(* Logix 5000 project; controller Seperator 1756-L85E rev 33.11; software revision 33.01; part 5 of 7 *)
(* tags used below, declared in another part *)
   batchstrng : STRING;
   bottle_clamp_out_delay : TIMER;
   bottle_clamp_out_delayF1 : TIMER;
   CAP_clamps_out_Delay : TIMER;
   Capper_Head_Sequencer : DINT;
   colours : STRING[3];
   Filler_Index_complete : BOOL;
   Filling : SFC_STEP;
   Filling_Nozzle_Down_Delay1 : TIMER;
   Filling_Nozzle_up_Delay1 : TIMER;
   Logix_Status : Logix_Status_FP;
   Qtr_Sec_PLs : TIMER;
   Random : AOI_SIM_RNG_Simple;

PROGRAM Capper_Heads   (* main routine Initialisation *)
VAR
   Alias_Head_Clamp_Pressure_SP : ALIAS FOR Head_Clamp_Pressure_SP;
   Bottle_Clamp_Pressure_actual : REAL := 10.799999;
   Cap_Pressure : REAL := 9.4;
   Head1_98_Percent_temperatureSP : REAL := 176.4;
   Head_Clamp_Pressure_SP : REAL := 90.0;
   Head_Down : BOOL;
   Head_Down_Stage1 : REAL := 18.0;
   Head_Down_Stage2 : REAL := 27.0;
   Head_Injection_Pressure_SP : REAL := 75.0;
   Head_Injection_Stage1 : REAL := 18.75;
   Head_Injection_Stage2 : REAL := 33.75;
   Head_Injector_out_delay : TIMER := (PRE := 2000);
   Head_moving_Down : BOOL := 1;
   Head_moving_Up : BOOL;
   Head_Up : BOOL;
   Head_up_delay : TIMER := (PRE := 2000);
   Pump_Running : BOOL := 1;
   Rotary_Moulder_Head_Name : STRING := 'Head 1'; {constant, access None}
   ScratchPad1 : REAL := 0.9;
   ScratchPad2 : REAL := 0.9;
   ScratchPad3 : REAL := 0.75;
   ScratchPad4 : REAL := 0.75;
   ScratchPad5 : REAL := 3.6;
   ScratchPad6 : REAL;
END_VAR

ROUTINE Head_Control   (* ladder *)
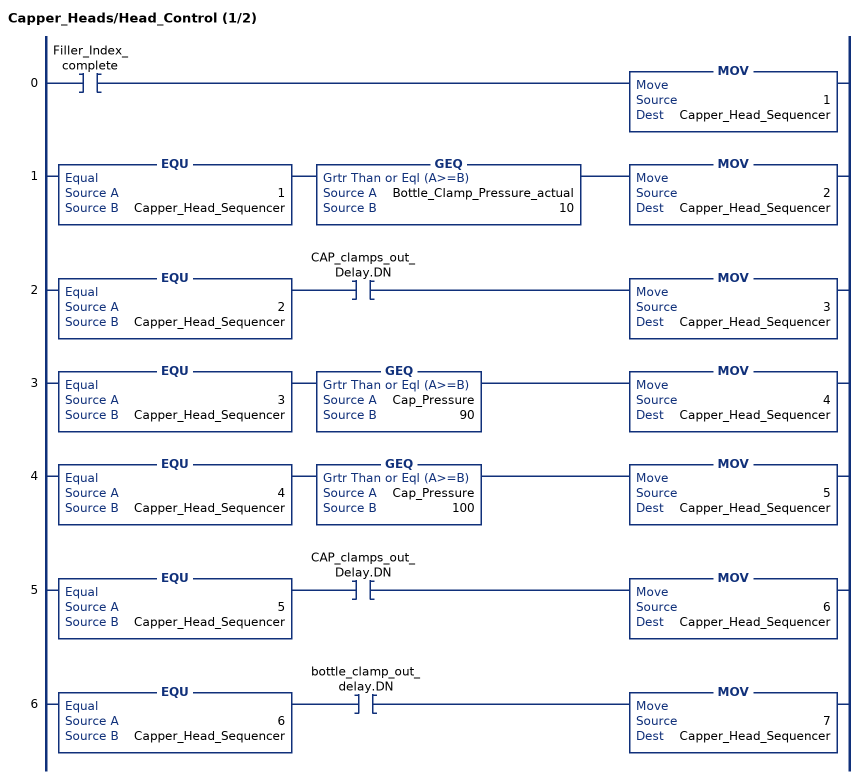
   0: XIC(Filler_Index_complete)MOV(1,Capper_Head_Sequencer);
   1: EQU(1,Capper_Head_Sequencer)GEQ(Bottle_Clamp_Pressure_actual,10)MOV(2,Capper_Head_Sequencer);
   2: EQU(2,Capper_Head_Sequencer)XIC(CAP_clamps_out_Delay.DN)MOV(3,Capper_Head_Sequencer);
   3: EQU(3,Capper_Head_Sequencer)GEQ(Cap_Pressure,90)MOV(4,Capper_Head_Sequencer);
   4: EQU(4,Capper_Head_Sequencer)GEQ(Cap_Pressure,100)MOV(5,Capper_Head_Sequencer);
   5: EQU(5,Capper_Head_Sequencer)XIC(CAP_clamps_out_Delay.DN)MOV(6,Capper_Head_Sequencer);
   6: EQU(6,Capper_Head_Sequencer)XIC(bottle_clamp_out_delay.DN)MOV(7,Capper_Head_Sequencer);
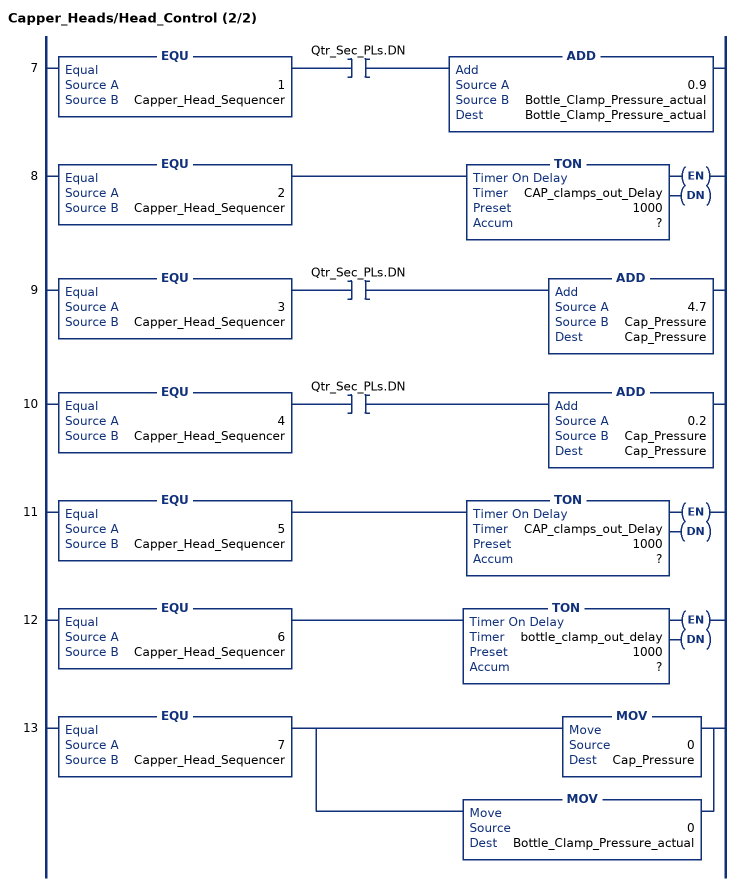
   7: EQU(1,Capper_Head_Sequencer)XIC(Qtr_Sec_PLs.DN)ADD(0.9,Bottle_Clamp_Pressure_actual,Bottle_Clamp_Pressure_actual);
   8: EQU(2,Capper_Head_Sequencer)TON(CAP_clamps_out_Delay,?,?);
   9: EQU(3,Capper_Head_Sequencer)XIC(Qtr_Sec_PLs.DN)ADD(4.7,Cap_Pressure,Cap_Pressure);
   10: EQU(4,Capper_Head_Sequencer)XIC(Qtr_Sec_PLs.DN)ADD(0.2,Cap_Pressure,Cap_Pressure);
   11: EQU(5,Capper_Head_Sequencer)TON(CAP_clamps_out_Delay,?,?);
   12: EQU(6,Capper_Head_Sequencer)TON(bottle_clamp_out_delay,?,?);
   13: EQU(7,Capper_Head_Sequencer)[MOV(0,Cap_Pressure) ,MOV(0,Bottle_Clamp_Pressure_actual) ];
END_ROUTINE

ROUTINE Head_HMI_Collation   (* ladder *)
END_ROUTINE

ROUTINE Initialisation   (* ladder *)
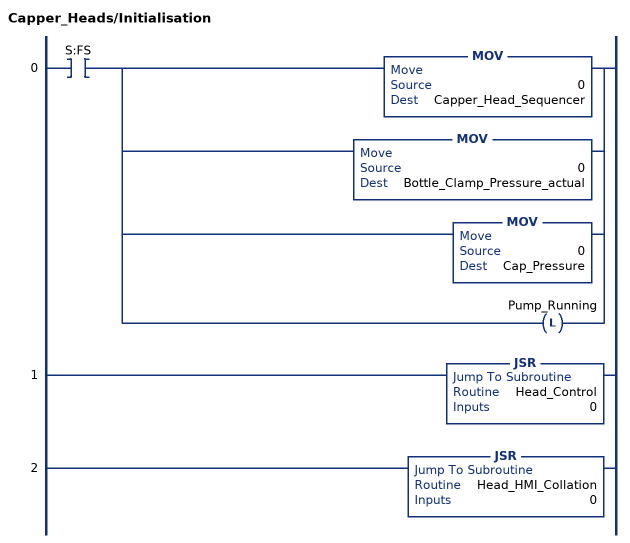
   0: XIC(S:FS)[MOV(0,Capper_Head_Sequencer) ,MOV(0,Bottle_Clamp_Pressure_actual) ,MOV(0,Cap_Pressure) ,OTL(Pump_Running) ];
   1: JSR(Head_Control,0);
   2: JSR(Head_HMI_Collation,0);
END_ROUTINE
END_PROGRAM

PROGRAM Controller_Fault   (* main routine Major_Controller_Fault *)

ROUTINE Major_Controller_Fault   (* ladder *)
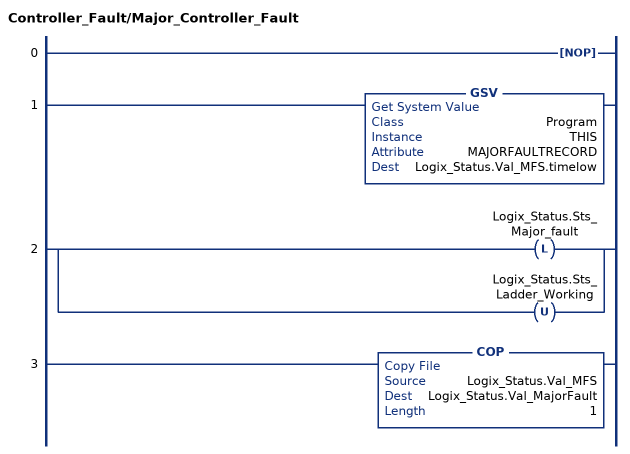
   0: NOP();
   1: GSV(Program,THIS,MAJORFAULTRECORD,Logix_Status.Val_MFS.timelow);
   2: [OTL(Logix_Status.Sts_Major_fault) ,OTU(Logix_Status.Sts_Ladder_Working) ];
   3: COP(Logix_Status.Val_MFS,Logix_Status.Val_MajorFault,1);
END_ROUTINE
END_PROGRAM

PROGRAM Filler   (* main routine Initialisation *)
VAR
   autoreset : TIMER := (PRE := 38913);
   autoresetpulse : BOOL;
   batchcountbase : DINT := 35000;
   batchcounter : DINT := 704;
   colourcounter : DINT := 2;
   Filler1_Heater_Tripped : ALARM_DIGITAL;
   Filler1_Hyd_Oil_Pressure_Low : ALARM_DIGITAL;
   Filler1_Hyd_Pump_Failure : ALARM_DIGITAL;
   Filler1_Index_Failure : ALARM_DIGITAL;
   Filler1_Overload : ALARM_DIGITAL;
   Filler_Efficiency_FTAE : BOOL[32];
   Filler_Fault_FTAE : BOOL[32];
   Filler_Heater_Tripped : BOOL;
   Filler_Hyd_Oil_Pressure_Low : BOOL;
   Filler_Hyd_Pump_Failure : BOOL;
   Filler_Index_Failure : BOOL;
   Filler_Overload : BOOL;
   Filler_Running : BOOL := 1;
   Filler_Warning_FTAE : BOOL[32];
   Index_Move : BOOL;
   Index_Move_Timer : TIMER := (PRE := 1000);
   m_slowperc_lim : REAL := 0.92;
   MetricsData : mtrcsdt := (PartId := 'Corner block', IdealCT := 23.7, GoodParts := 30066, ScrapParts := 5250, TotalParts := 35316, Running := 1, Monitored_Availability := 1, Machine_State := 1, BatchID := 'Batch ID 35704', Colour := 'White');
   mset_badperc : REAL := 0.07;   // Bad percentage valid: 1.0 - mset_goodperc
   mset_fltfudge : REAL := 0.93;   // fault distribution fudge factor do not change
   mset_fltoffset : DINT := 2;   // fault distribution offset do not change
   mset_goodperc : REAL := 0.85;   // Good percentage valid: 0.51 - 0.99
   mset_wrnfudge : REAL := 0.02;   // warning distribution fudge factor do not change
   mset_wrnoffset : DINT := 2;   // warning distribution offset do not change
   oneshots : DINT;
   tempDINT : DINT := 16;
   tempstring : STRING := '35704';
END_VAR

ROUTINE Filler_Alarms   (* ladder *)
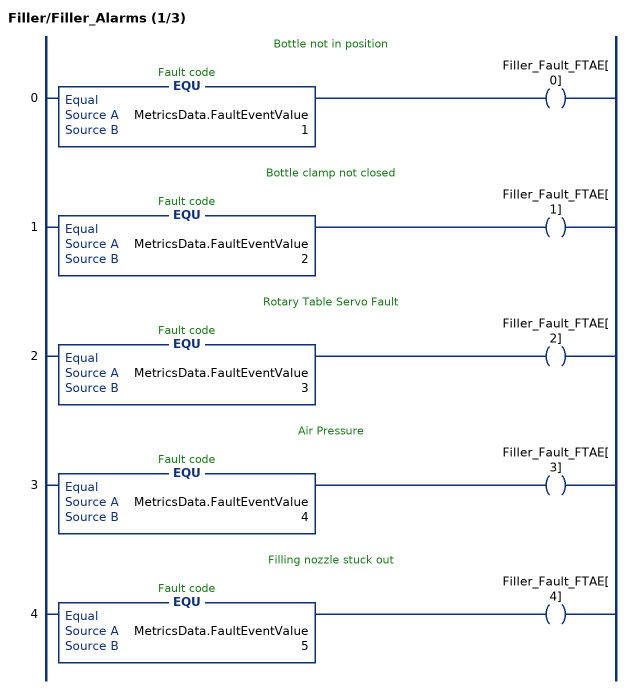
   // Bottle not in position
   0: EQU(MetricsData.FaultEventValue,1)OTE(Filler_Fault_FTAE[0]);
   // Bottle clamp not closed
   1: EQU(MetricsData.FaultEventValue,2)OTE(Filler_Fault_FTAE[1]);
   // Rotary Table Servo Fault
   2: EQU(MetricsData.FaultEventValue,3)OTE(Filler_Fault_FTAE[2]);
   // Air Pressure
   3: EQU(MetricsData.FaultEventValue,4)OTE(Filler_Fault_FTAE[3]);
   // Filling nozzle stuck out
   4: EQU(MetricsData.FaultEventValue,5)OTE(Filler_Fault_FTAE[4]);
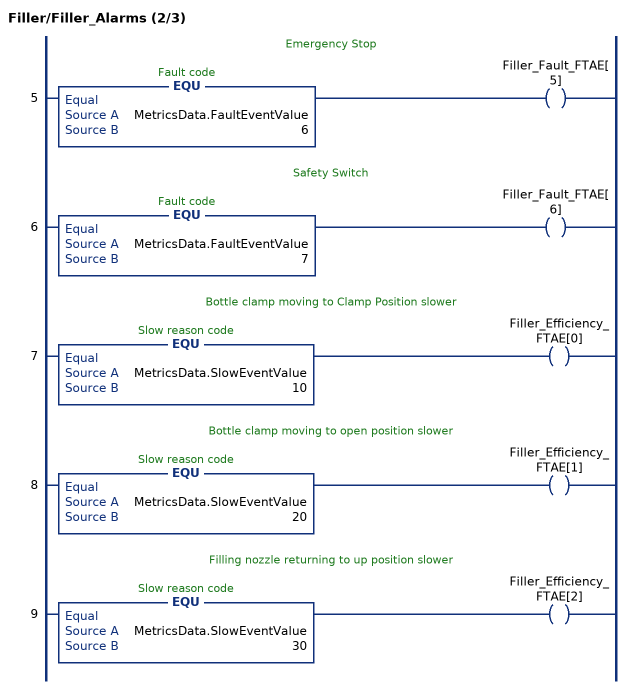
   // Emergency Stop
   5: EQU(MetricsData.FaultEventValue,6)OTE(Filler_Fault_FTAE[5]);
   // Safety Switch
   6: EQU(MetricsData.FaultEventValue,7)OTE(Filler_Fault_FTAE[6]);
   // Bottle clamp moving to Clamp Position slower
   7: EQU(MetricsData.SlowEventValue,10)OTE(Filler_Efficiency_FTAE[0]);
   // Bottle clamp moving to open position slower
   8: EQU(MetricsData.SlowEventValue,20)OTE(Filler_Efficiency_FTAE[1]);
   // Filling nozzle returning to up position slower
   9: EQU(MetricsData.SlowEventValue,30)OTE(Filler_Efficiency_FTAE[2]);
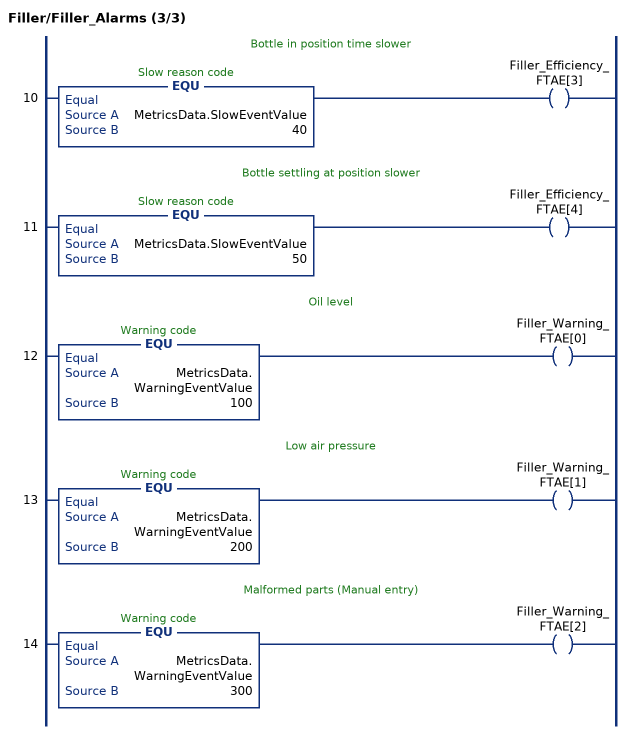
   // Bottle in position time slower
   10: EQU(MetricsData.SlowEventValue,40)OTE(Filler_Efficiency_FTAE[3]);
   // Bottle settling at position slower
   11: EQU(MetricsData.SlowEventValue,50)OTE(Filler_Efficiency_FTAE[4]);
   // Oil level
   12: EQU(MetricsData.WarningEventValue,100)OTE(Filler_Warning_FTAE[0]);
   // Low air pressure
   13: EQU(MetricsData.WarningEventValue,200)OTE(Filler_Warning_FTAE[1]);
   // Malformed parts (Manual entry)
   14: EQU(MetricsData.WarningEventValue,300)OTE(Filler_Warning_FTAE[2]);
END_ROUTINE

ROUTINE Index_Control   (* ladder *)
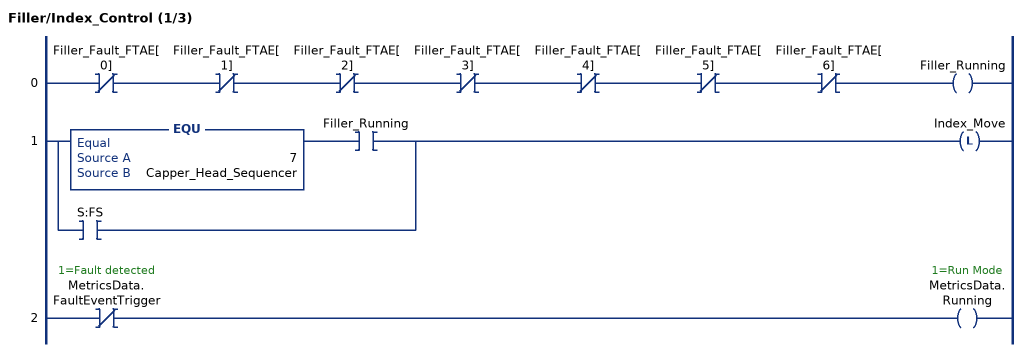
   0: XIO(Filler_Fault_FTAE[0])XIO(Filler_Fault_FTAE[1])XIO(Filler_Fault_FTAE[2])XIO(Filler_Fault_FTAE[3])XIO(Filler_Fault_FTAE[4])XIO(Filler_Fault_FTAE[5])XIO(Filler_Fault_FTAE[6])OTE(Filler_Running);
   1: [EQU(7,Capper_Head_Sequencer) XIC(Filler_Running) ,XIC(S:FS) ]OTL(Index_Move);
   2: XIO(MetricsData.FaultEventTrigger)OTE(MetricsData.Running);
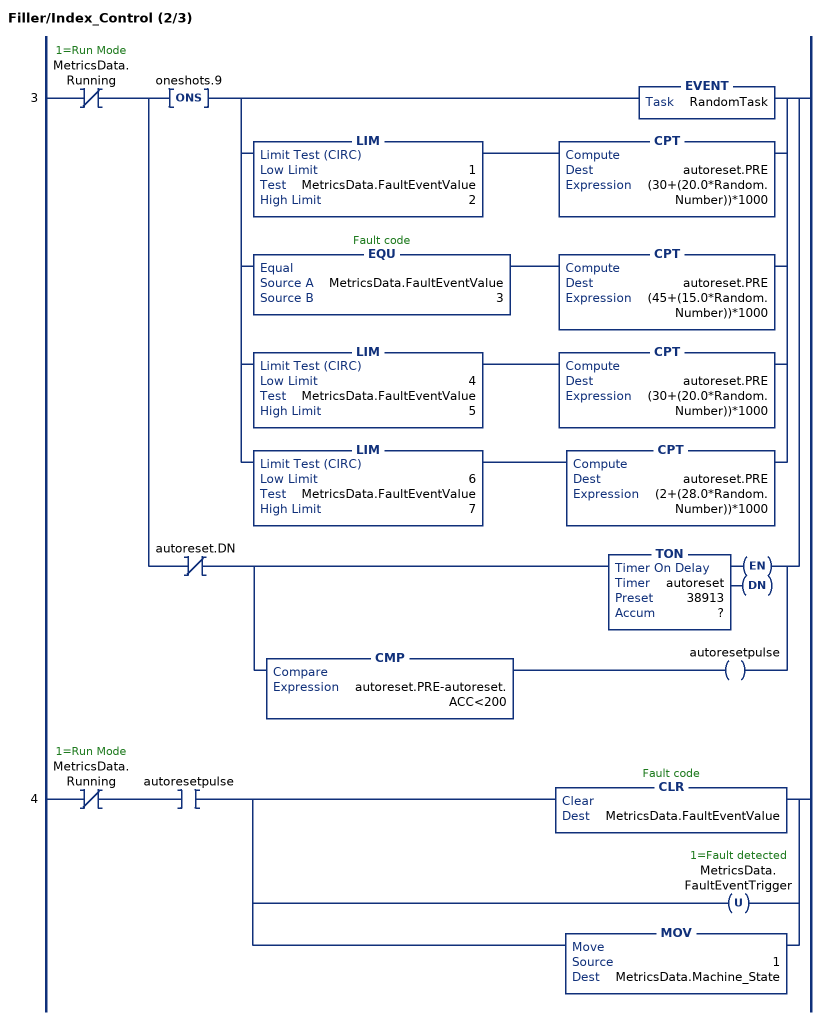
   3: XIO(MetricsData.Running)[ONS(oneshots.9) [EVENT(RandomTask) ,LIM(1,MetricsData.FaultEventValue,2) CPT(autoreset.PRE,(30+(20.0*Random.Number))*1000) ,EQU(MetricsData.FaultEventValue,3) CPT(autoreset.PRE,(45+(15.0*Random.Number))*1000) ,LIM(4,MetricsData.FaultEventValue,5) CPT(autoreset.PRE,(30+(20.0*Random.Number))*1000) ,LIM(6,MetricsData.FaultEventValue,7) CPT(autoreset.PRE,(2+(28.0*Random.Number))*1000) ] ,XIO(autoreset.DN) [TON(autoreset,?,?) ,CMP(autoreset.PRE-autoreset.ACC<200) OTE(autoresetpulse) ] ];
   4: XIO(MetricsData.Running)XIC(autoresetpulse)[CLR(MetricsData.FaultEventValue) ,OTU(MetricsData.FaultEventTrigger) ,MOV(1,MetricsData.Machine_State) ];
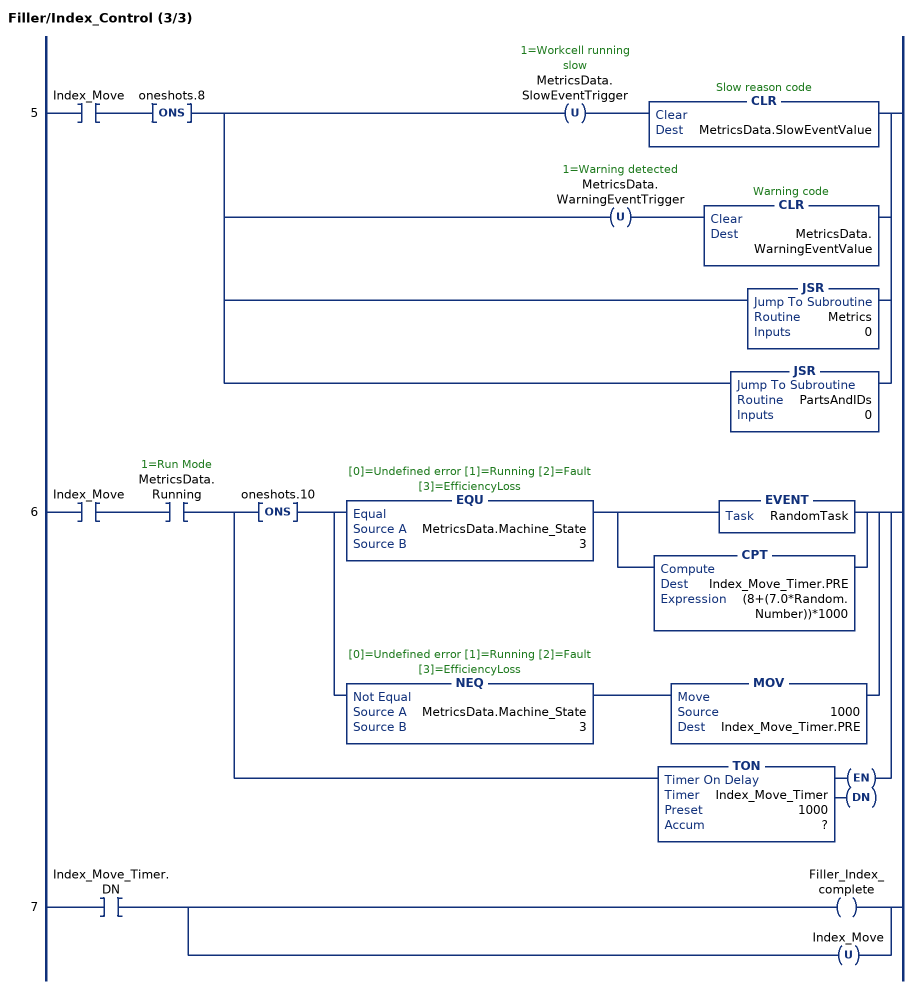
   5: XIC(Index_Move)ONS(oneshots.8)[OTU(MetricsData.SlowEventTrigger) CLR(MetricsData.SlowEventValue) ,OTU(MetricsData.WarningEventTrigger) CLR(MetricsData.WarningEventValue) ,JSR(Metrics,0) ,JSR(PartsAndIDs,0) ];
   6: XIC(Index_Move)XIC(MetricsData.Running)[ONS(oneshots.10) [EQU(MetricsData.Machine_State,3) [EVENT(RandomTask) ,CPT(Index_Move_Timer.PRE,(8+(7.0*Random.Number))*1000) ] ,NEQ(MetricsData.Machine_State,3) MOV(1000,Index_Move_Timer.PRE) ] ,TON(Index_Move_Timer,?,?) ];
   7: XIC(Index_Move_Timer.DN)[OTE(Filler_Index_complete) ,OTU(Index_Move) ];
END_ROUTINE

ROUTINE Initialisation   (* ladder *)
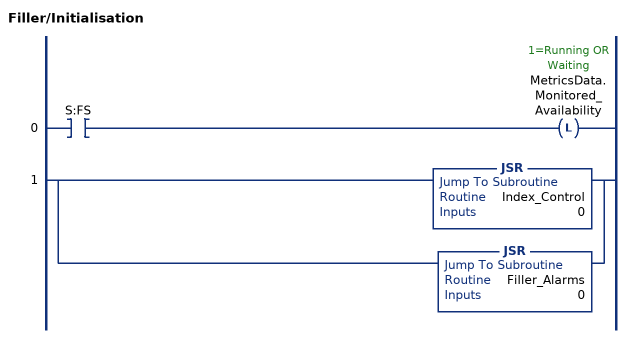
   0: XIC(S:FS)OTL(MetricsData.Monitored_Availability);
   1: [JSR(Index_Control,0) ,JSR(Filler_Alarms,0) ];
END_ROUTINE

ROUTINE Metrics   (* ladder *)
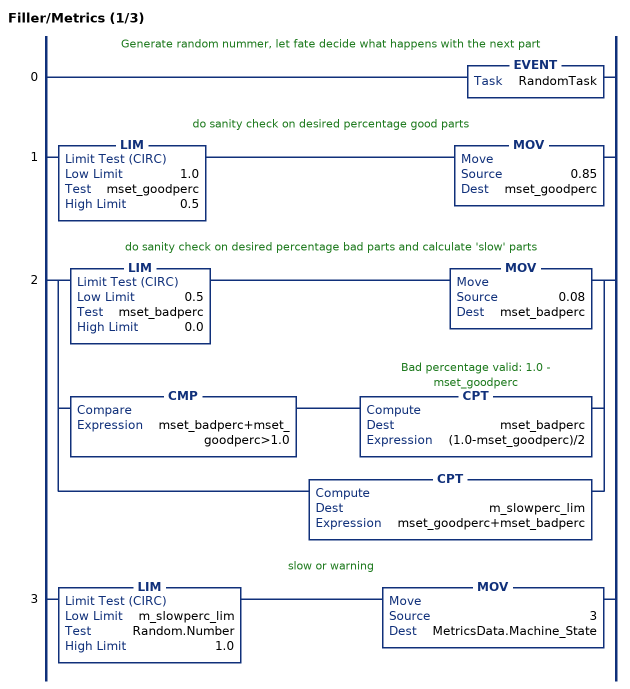
   // Generate random nummer, let fate decide what happens with the next part
   0: EVENT(RandomTask);
   // do sanity check on desired percentage good parts
   1: LIM(1.0,mset_goodperc,0.5)MOV(0.85,mset_goodperc);
   // do sanity check on desired percentage bad parts and calculate 'slow' parts
   2: [LIM(0.5,mset_badperc,0.0) MOV(0.08,mset_badperc) ,CMP(mset_badperc+mset_goodperc>1.0) CPT(mset_badperc,(1.0-mset_goodperc)/2) ,CPT(m_slowperc_lim,mset_goodperc+mset_badperc) ];
   // slow or warning
   3: LIM(m_slowperc_lim,Random.Number,1.0)MOV(3,MetricsData.Machine_State);
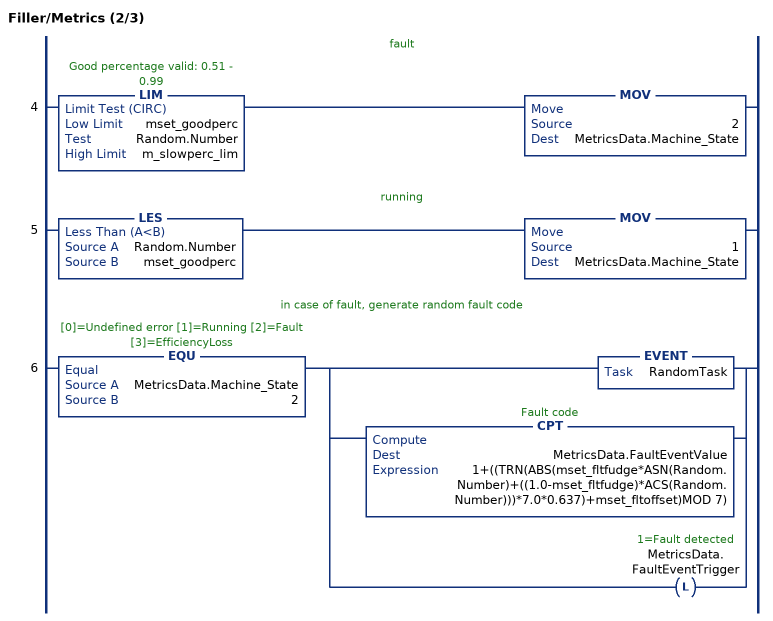
   // fault
   4: LIM(mset_goodperc,Random.Number,m_slowperc_lim)MOV(2,MetricsData.Machine_State);
   // running
   5: LES(Random.Number,mset_goodperc)MOV(1,MetricsData.Machine_State);
   // in case of fault, generate random fault code
   6: EQU(MetricsData.Machine_State,2)[EVENT(RandomTask) ,CPT(MetricsData.FaultEventValue,1+((TRN(ABS(mset_fltfudge*ASN(Random.Number)+((1.0-mset_fltfudge)*ACS(Random.Number)))*7.0*0.637)+mset_fltoffset)MOD 7)) ,OTL(MetricsData.FaultEventTrigger) ];
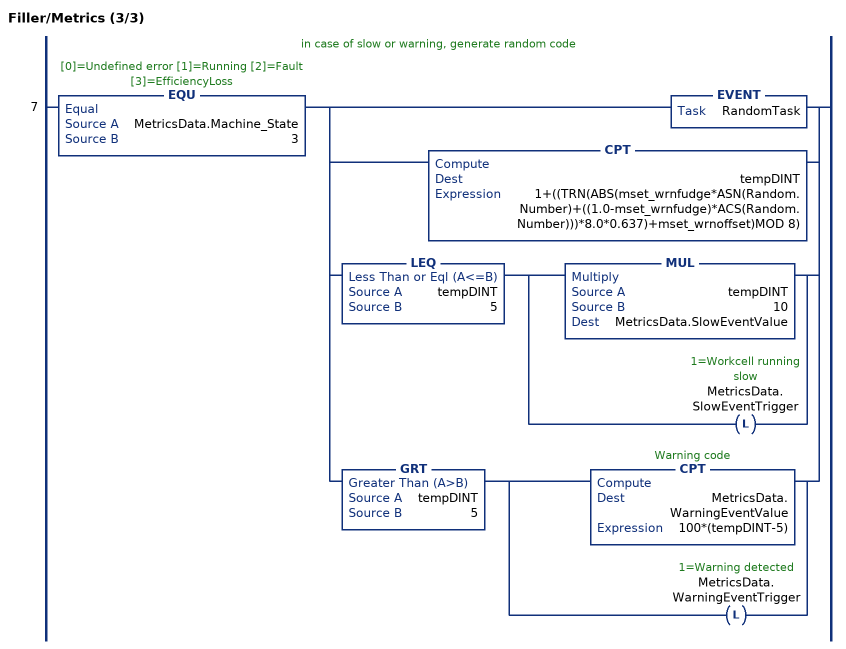
   // in case of slow or warning, generate random code
   7: EQU(MetricsData.Machine_State,3)[EVENT(RandomTask) ,CPT(tempDINT,1+((TRN(ABS(mset_wrnfudge*ASN(Random.Number)+((1.0-mset_wrnfudge)*ACS(Random.Number)))*8.0*0.637)+mset_wrnoffset)MOD 8)) ,LEQ(tempDINT,5) [MUL(tempDINT,10,MetricsData.SlowEventValue) ,OTL(MetricsData.SlowEventTrigger) ] ,GRT(tempDINT,5) [CPT(MetricsData.WarningEventValue,100*(tempDINT-5)) ,OTL(MetricsData.WarningEventTrigger) ] ];
END_ROUTINE

ROUTINE PartsAndIDs   (* ladder *)
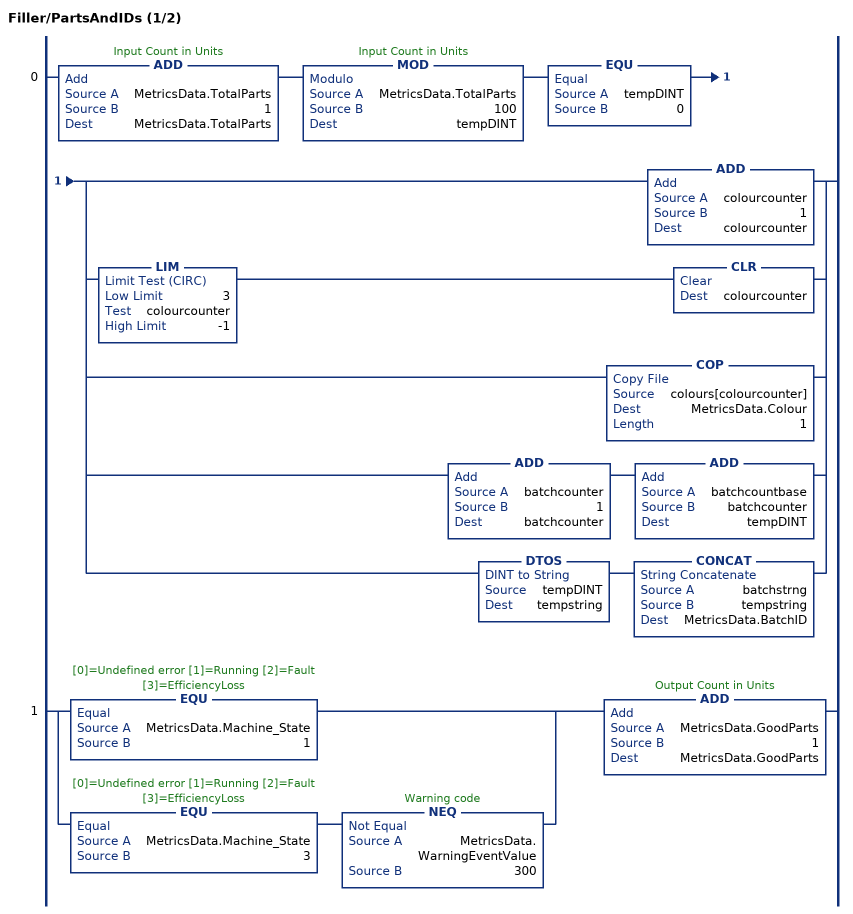
   0: ADD(MetricsData.TotalParts,1,MetricsData.TotalParts)MOD(MetricsData.TotalParts,100,tempDINT)EQU(tempDINT,0)[ADD(colourcounter,1,colourcounter) ,LIM(3,colourcounter,-1) CLR(colourcounter) ,COP(colours[colourcounter],MetricsData.Colour,1) ,ADD(batchcounter,1,batchcounter) ADD(batchcountbase,batchcounter,tempDINT) ,DTOS(tempDINT,tempstring) CONCAT(batchstrng,tempstring,MetricsData.BatchID) ];
   1: [EQU(MetricsData.Machine_State,1) ,EQU(MetricsData.Machine_State,3) NEQ(MetricsData.WarningEventValue,300) ]ADD(MetricsData.GoodParts,1,MetricsData.GoodParts);
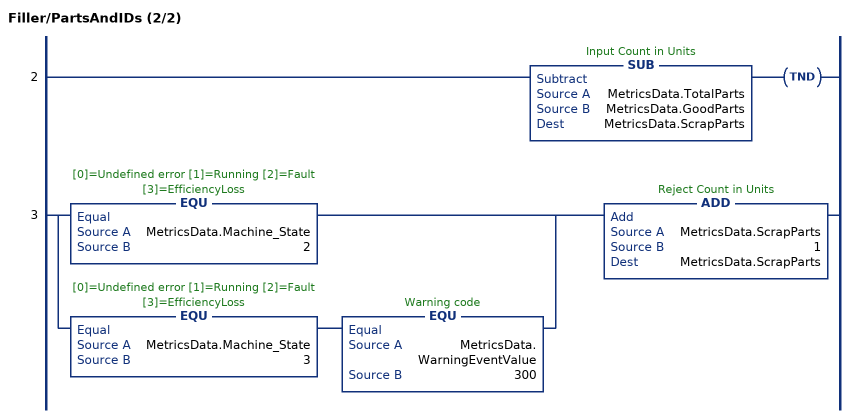
   2: SUB(MetricsData.TotalParts,MetricsData.GoodParts,MetricsData.ScrapParts)TND();
   3: [EQU(MetricsData.Machine_State,2) ,EQU(MetricsData.Machine_State,3) EQU(MetricsData.WarningEventValue,300) ]ADD(MetricsData.ScrapParts,1,MetricsData.ScrapParts);
END_ROUTINE
END_PROGRAM

PROGRAM Filler_Heads1   (* main routine Initialisation *)
VAR
   Alias_Head_Clamp_Pressure_SP_1 : ALIAS FOR Head_Clamp_Pressure_SP_1;
   Bottle_Clamp_Pressure_actual_1 : REAL := 10.799999;
   Bottle_Clamp_Pressure_SP_1 : REAL := 10.0;
   Bottle_level_actual_1 : REAL := 9.4;
   Bottle_Slow_Fill_SP_1 : REAL := 90.0;
   Bottle_Stop_Fill_SP_1 : REAL := 100.0;
   Filling_Head_Sequencer_1 : DINT := 3;
   Head1_98_Percent_temperatureSP_1 : REAL := 176.4;
   Head_Clamp_Pressure_SP_1 : REAL := 90.0;
   Head_Down_1 : BOOL;
   Head_Down_Stage1_1 : REAL := 18.0;
   Head_Down_Stage2_1 : REAL := 27.0;
   Head_Injection_Pressure_SP_1 : REAL := 75.0;
   Head_Injection_Stage1_1 : REAL := 18.75;
   Head_Injection_Stage2_1 : REAL := 33.75;
   Head_Injector_out_delay_1 : TIMER := (PRE := 2000);
   Head_moving_Down_1 : BOOL := 1;
   Head_moving_Up_1 : BOOL;
   Head_Up_1 : BOOL;
   Head_up_delay_1 : TIMER := (PRE := 2000);
   Pump_Running_1 : BOOL := 1;
   Rotary_Moulder_Head_Name_1 : STRING := 'Head 1'; {constant, access None}
   ScratchPad1_1 : REAL := 0.9;
   ScratchPad2_1 : REAL := 0.9;
   ScratchPad3_1 : REAL := 0.75;
   ScratchPad4_1 : REAL := 0.75;
   ScratchPad5_1 : REAL := 3.6;
   ScratchPad6_1 : REAL;
END_VAR

ROUTINE Head_Control   (* ladder *)
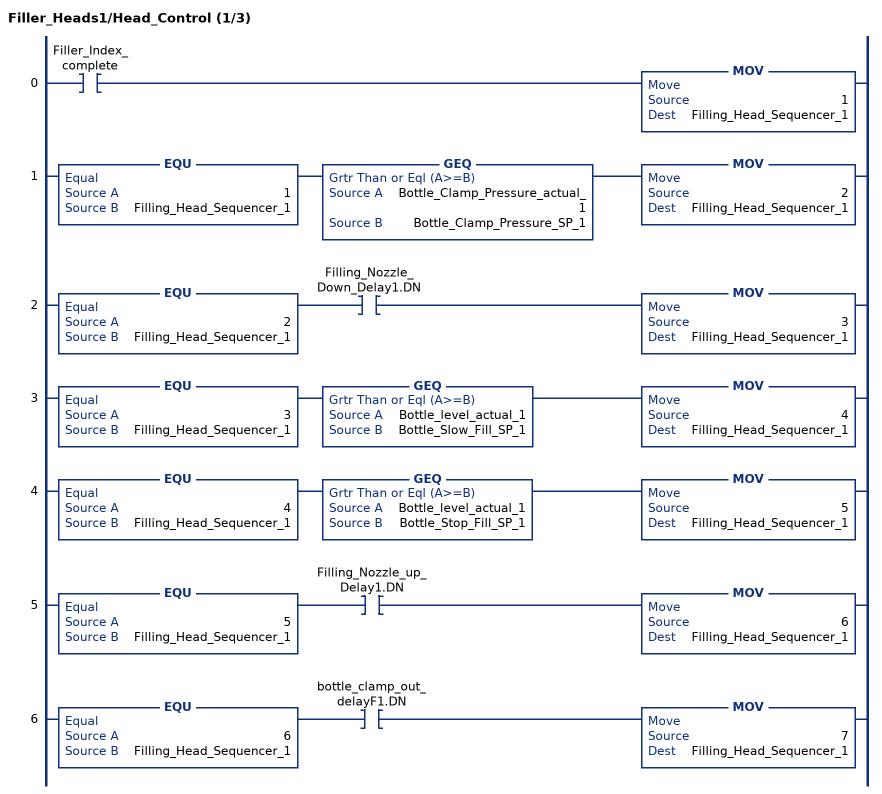
   0: XIC(Filler_Index_complete)MOV(1,Filling_Head_Sequencer_1);
   1: EQU(1,Filling_Head_Sequencer_1)GEQ(Bottle_Clamp_Pressure_actual_1,Bottle_Clamp_Pressure_SP_1)MOV(2,Filling_Head_Sequencer_1);
   2: EQU(2,Filling_Head_Sequencer_1)XIC(Filling_Nozzle_Down_Delay1.DN)MOV(3,Filling_Head_Sequencer_1);
   3: EQU(3,Filling_Head_Sequencer_1)GEQ(Bottle_level_actual_1,Bottle_Slow_Fill_SP_1)MOV(4,Filling_Head_Sequencer_1);
   4: EQU(4,Filling_Head_Sequencer_1)GEQ(Bottle_level_actual_1,Bottle_Stop_Fill_SP_1)MOV(5,Filling_Head_Sequencer_1);
   5: EQU(5,Filling_Head_Sequencer_1)XIC(Filling_Nozzle_up_Delay1.DN)MOV(6,Filling_Head_Sequencer_1);
   6: EQU(6,Filling_Head_Sequencer_1)XIC(bottle_clamp_out_delayF1.DN)MOV(7,Filling_Head_Sequencer_1);
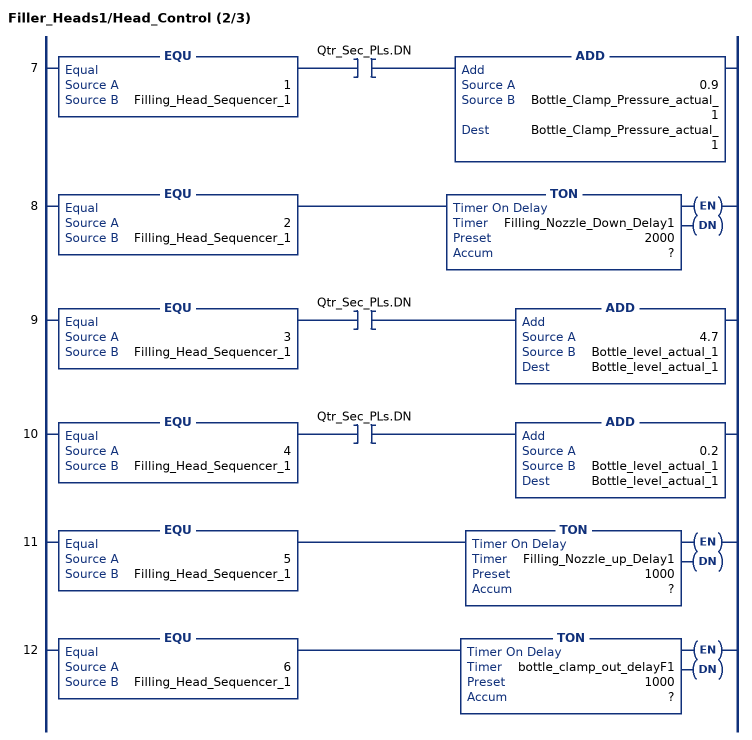
   7: EQU(1,Filling_Head_Sequencer_1)XIC(Qtr_Sec_PLs.DN)ADD(0.9,Bottle_Clamp_Pressure_actual_1,Bottle_Clamp_Pressure_actual_1);
   8: EQU(2,Filling_Head_Sequencer_1)TON(Filling_Nozzle_Down_Delay1,?,?);
   9: EQU(3,Filling_Head_Sequencer_1)XIC(Qtr_Sec_PLs.DN)ADD(4.7,Bottle_level_actual_1,Bottle_level_actual_1);
   10: EQU(4,Filling_Head_Sequencer_1)XIC(Qtr_Sec_PLs.DN)ADD(0.2,Bottle_level_actual_1,Bottle_level_actual_1);
   11: EQU(5,Filling_Head_Sequencer_1)TON(Filling_Nozzle_up_Delay1,?,?);
   12: EQU(6,Filling_Head_Sequencer_1)TON(bottle_clamp_out_delayF1,?,?);
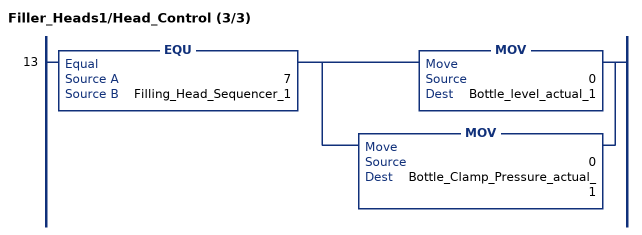
   13: EQU(7,Filling_Head_Sequencer_1)[MOV(0,Bottle_level_actual_1) ,MOV(0,Bottle_Clamp_Pressure_actual_1) ];
END_ROUTINE
